REGION Network 5: State 2 = Valves Control
   RUNG wire#powerrail
      Contact( #RUNNING )
      { S7_Templates := "SrcType := Int" } GE_Contact(in1 := #STATE, in2 := 2)
      wire#w1
      { S7_Templates := "SrcType := Int" } LT_Contact(in1 := #STATE, in2 := 6)
      Coil( #OPN_AV )
   END_RUNG
   RUNG wire#w1
      { S7_Templates := "SrcType := Int" } LT_Contact(in1 := #STATE, in2 := 4)
      Coil( #OPN_FV1 )
   END_RUNG
   RUNG wire#w1
      { S7_Templates := "SrcType := Int" } LT_Contact(in1 := #STATE, in2 := 5)
      wire#w2
      Coil( #OPN_3W_FV2 )
   END_RUNG
   RUNG wire#w1
      { S7_Templates := "SrcType := Int" } GE_Contact(in1 := #STATE, in2 := 7)
      { S7_Templates := "SrcType := Int" } LE_Contact(in1 := #STATE, in2 := 8)
   END_RUNG wire#w2
   // the same network as SCL:
   #_w1 := #RUNNING AND (#STATE >= 2);
   #OPN_AV := #_w1 AND (#STATE < 6);
   #OPN_FV1 := #_w1 AND (#STATE < 4);
   #OPN_3W_FV2 := #_w1 AND ((#STATE < 5) OR ((#STATE >= 7) AND (#STATE <= 8)));
END_REGION

REGION Network 6: Into State 3
   RUNG wire#powerrail
      Contact( #RUNNING )
      { S7_Templates := "SrcType := Int" } EQ_Contact(in1 := #STATE, in2 := 2)
      Contact( #AV_Q )
      Contact( #FV1_Q )
      Contact( #FV2_3W_Q )
      Move(in := 3, out1 => #STATE)
   END_RUNG
   // the same network as SCL:
   IF #RUNNING AND (#STATE = 2) AND #AV_Q AND #FV1_Q AND #FV2_3W_Q THEN #STATE := 3; END_IF;
END_REGION

REGION Network 7: State 3 = Purge Active
   RUNG wire#powerrail
      Contact( #RUNNING )
      { S7_Templates := "SrcType := Int" } GE_Contact(in1 := #STATE, in2 := 3)
      { S7_Templates := "SrcType := Int" } LE_Contact(in1 := #STATE, in2 := 8)
      wire#w1
      Coil( #PRG_ACTV )
   END_RUNG
   RUNG wire#w1
      Coil( #ACTIVE )
   END_RUNG
   // the same network as SCL:
   #PRG_ACTV := #RUNNING AND (#STATE >= 3) AND (#STATE <= 8);
   #ACTIVE := #PRG_ACTV;
END_REGION

REGION Network 8: Into State 4
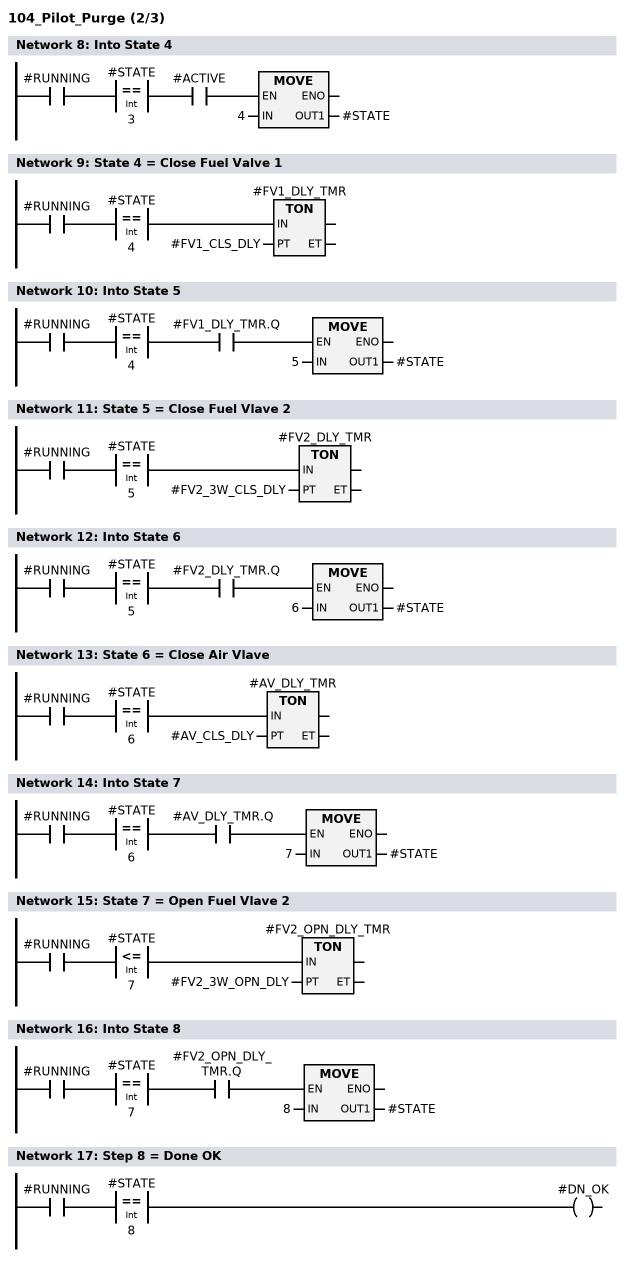
   RUNG wire#powerrail
      Contact( #RUNNING )
      { S7_Templates := "SrcType := Int" } EQ_Contact(in1 := #STATE, in2 := 3)
      Contact( #ACTIVE )
      Move(in := 4, out1 => #STATE)
   END_RUNG
   // the same network as SCL:
   IF #RUNNING AND (#STATE = 3) AND #ACTIVE THEN #STATE := 4; END_IF;
END_REGION

REGION Network 9: State 4 = Close Fuel Valve 1
   #FV1_DLY_TMR(IN := #RUNNING AND (#STATE = 4), PT := #FV1_CLS_DLY);   // TON
END_REGION

REGION Network 10: Into State 5
   RUNG wire#powerrail
      Contact( #RUNNING )
      { S7_Templates := "SrcType := Int" } EQ_Contact(in1 := #STATE, in2 := 4)
      Contact( #FV1_DLY_TMR.Q )
      Move(in := 5, out1 => #STATE)
   END_RUNG
   // the same network as SCL:
   IF #RUNNING AND (#STATE = 4) AND #FV1_DLY_TMR.Q THEN #STATE := 5; END_IF;
END_REGION

REGION Network 11: State 5 = Close Fuel Vlave 2
   #FV2_DLY_TMR(IN := #RUNNING AND (#STATE = 5), PT := #FV2_3W_CLS_DLY);   // TON
END_REGION

REGION Network 12: Into State 6
   RUNG wire#powerrail
      Contact( #RUNNING )
      { S7_Templates := "SrcType := Int" } EQ_Contact(in1 := #STATE, in2 := 5)
      Contact( #FV2_DLY_TMR.Q )
      Move(in := 6, out1 => #STATE)
   END_RUNG
   // the same network as SCL:
   IF #RUNNING AND (#STATE = 5) AND #FV2_DLY_TMR.Q THEN #STATE := 6; END_IF;
END_REGION

REGION Network 13: State 6 = Close Air Vlave
   #AV_DLY_TMR(IN := #RUNNING AND (#STATE = 6), PT := #AV_CLS_DLY);   // TON
END_REGION

REGION Network 14: Into State 7
   RUNG wire#powerrail
      Contact( #RUNNING )
      { S7_Templates := "SrcType := Int" } EQ_Contact(in1 := #STATE, in2 := 6)
      Contact( #AV_DLY_TMR.Q )
      Move(in := 7, out1 => #STATE)
   END_RUNG
   // the same network as SCL:
   IF #RUNNING AND (#STATE = 6) AND #AV_DLY_TMR.Q THEN #STATE := 7; END_IF;
END_REGION

REGION Network 15: State 7 = Open Fuel Vlave 2
   #FV2_OPN_DLY_TMR(IN := #RUNNING AND (#STATE <= 7), PT := #FV2_3W_OPN_DLY);   // TON
END_REGION

REGION Network 16: Into State 8
   RUNG wire#powerrail
      Contact( #RUNNING )
      { S7_Templates := "SrcType := Int" } EQ_Contact(in1 := #STATE, in2 := 7)
      Contact( #FV2_OPN_DLY_TMR.Q )
      Move(in := 8, out1 => #STATE)
   END_RUNG
   // the same network as SCL:
   IF #RUNNING AND (#STATE = 7) AND #FV2_OPN_DLY_TMR.Q THEN #STATE := 8; END_IF;
END_REGION

REGION Network 17: Step 8 = Done OK
   RUNG wire#powerrail
      Contact( #RUNNING )
      { S7_Templates := "SrcType := Int" } EQ_Contact(in1 := #STATE, in2 := 8)
      Coil( #DN_OK )
   END_RUNG
   // the same network as SCL:
   #DN_OK := #RUNNING AND (#STATE = 8);
END_REGION

REGION Network 18: Maximum Sequence Run Time
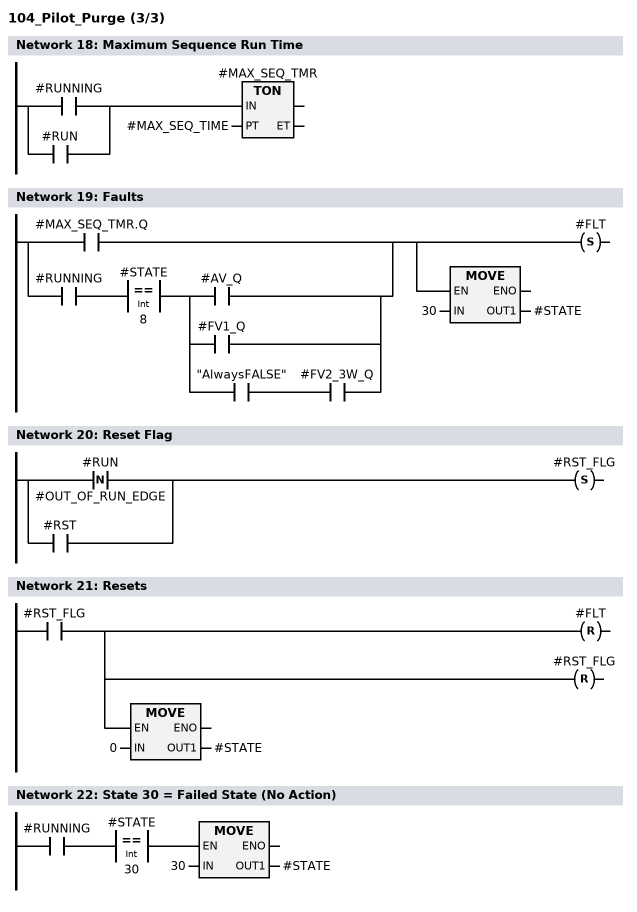
   #MAX_SEQ_TMR(IN := #RUNNING OR #RUN, PT := #MAX_SEQ_TIME);   // TON
END_REGION

REGION Network 19: Faults
   RUNG wire#powerrail
      Contact( #MAX_SEQ_TMR.Q )
      wire#w1
      S_Coil( #FLT )
   END_RUNG
   RUNG wire#powerrail
      Contact( #RUNNING )
      { S7_Templates := "SrcType := Int" } EQ_Contact(in1 := #STATE, in2 := 8)
      wire#w2
      Contact( #AV_Q )
   END_RUNG wire#w1
   RUNG wire#w2
      Contact( #FV1_Q )
   END_RUNG wire#w1
   RUNG wire#w2
      Contact( "AlwaysFALSE" )
      Contact( #FV2_3W_Q )
   END_RUNG wire#w1
   RUNG wire#w1
      Move(in := 30, out1 => #STATE)
   END_RUNG
   // the same network as SCL:
   IF #MAX_SEQ_TMR.Q OR (#RUNNING AND (#STATE = 8) AND (#AV_Q OR #FV1_Q OR ("AlwaysFALSE" AND #FV2_3W_Q))) THEN
       #FLT := TRUE;
       #STATE := 30;
   END_IF;
END_REGION

REGION Network 20: Reset Flag
   RUNG wire#powerrail
      N_Contact(operand := #RUN, bit := #OUT_OF_RUN_EDGE)
      wire#w1
      S_Coil( #RST_FLG )
   END_RUNG
   RUNG wire#powerrail
      Contact( #RST )
   END_RUNG wire#w1
   // the same network as SCL:
   #_w1 := NOT #RUN AND #OUT_OF_RUN_EDGE;   // falling edge of #RUN
   #OUT_OF_RUN_EDGE := #RUN;
   IF #_w1 OR #RST THEN #RST_FLG := TRUE; END_IF;
END_REGION

REGION Network 21: Resets
   RUNG wire#powerrail
      Contact( #RST_FLG )
      wire#w1
      R_Coil( #FLT )
   END_RUNG
   RUNG wire#w1
      R_Coil( #RST_FLG )
   END_RUNG
   RUNG wire#w1
      Move(in := 0, out1 => #STATE)
   END_RUNG
   // the same network as SCL:
   IF #RST_FLG THEN #FLT := FALSE; END_IF;
   #_w1 := #RST_FLG;
   IF #_w1 THEN
       #RST_FLG := FALSE;
       #STATE := 0;
   END_IF;
END_REGION

REGION Network 22: State 30 = Failed State (No Action)
   RUNG wire#powerrail
      Contact( #RUNNING )
      { S7_Templates := "SrcType := Int" } EQ_Contact(in1 := #STATE, in2 := 30)
      Move(in := 30, out1 => #STATE)
   END_RUNG
   // the same network as SCL:
   IF #RUNNING AND (#STATE = 30) THEN #STATE := 30; END_IF;
END_REGION
END_FUNCTION_BLOCK

FUNCTION_BLOCK "Evolving Setpoint"   // FB105, LAD
{ S7_Optimized_Access := 'TRUE' }
VERSION : 0.1
   VAR_INPUT
      Enable : Bool;
      Value : Real;
      Setpoint : Real;
      Gain : Real;
      Level_High : Real;
      Level_Low : Real;
   END_VAR
   VAR_OUTPUT
      Gain_Derived : Real;
      LevelBetter : Bool;
   END_VAR
   VAR
      "OFF Time" : TON_TIME;
      "On Time" : TON_TIME;
      Aux : Struct
         Aux_Derived : Bool;
         AuxSenzorDerivata1 : Real;
         AuxSenzorDerivata2 : Real;
         AuxSenzorDerivata11 : Real;
         AuxSenzorDerivata12 : Real;
         Puls_1 : Bool;
         Puls_2 : Bool;
         Puls_3 : Bool;
         Puls_4 : Bool;
         Gain_1 : Real;
      END_STRUCT;
      "Delay TOF" : TOF_TIME;
      "LevelBetter Delay" : TOF_TIME;
      "LevelBetter Prolong" : TOF_TIME;
   END_VAR
   VAR_TEMP   // added for the SCL form of the ladder/FBD networks
      _w1 : Bool;
      _w2 : Bool;
      _w3 : Bool;
      _w4 : Bool;
      _w5 : Bool;
      _w6 : Bool;
   END_VAR
BEGIN

REGION Network 1: Calcul derivata
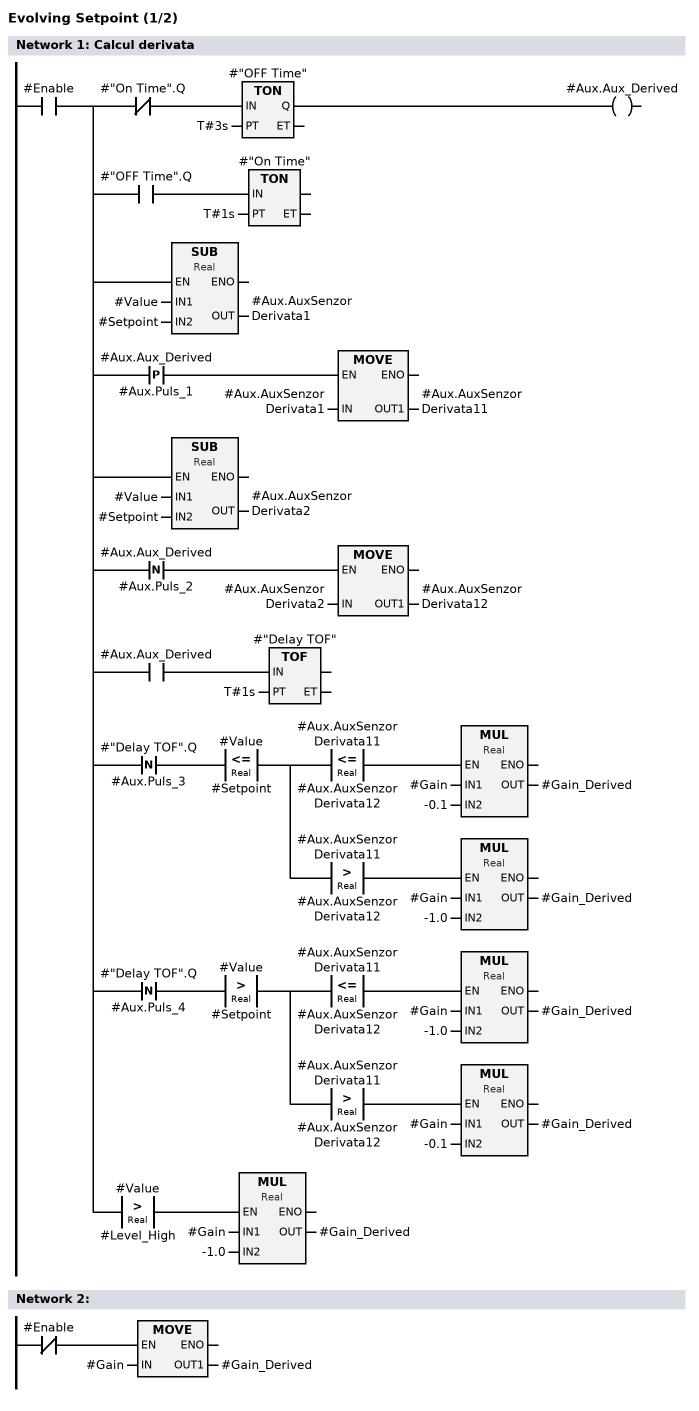
   #"OFF Time"(IN := #Enable AND NOT #"On Time".Q, PT := T#3s);   // TON
   #Aux.Aux_Derived := #"OFF Time".Q;
   #"On Time"(IN := #Enable AND #"OFF Time".Q, PT := T#1s);   // TON
   IF #Enable THEN #Aux.AuxSenzorDerivata1 := #Value - #Setpoint; END_IF;
   #_w1 := #Enable AND #Aux.Aux_Derived AND NOT #Aux.Puls_1;   // rising edge of #Aux.Aux_Derived
   #Aux.Puls_1 := #Aux.Aux_Derived;
   IF #_w1 THEN #Aux.AuxSenzorDerivata11 := #Aux.AuxSenzorDerivata1; END_IF;
   IF #Enable THEN #Aux.AuxSenzorDerivata2 := #Value - #Setpoint; END_IF;
   #_w2 := #Enable AND NOT #Aux.Aux_Derived AND #Aux.Puls_2;   // falling edge of #Aux.Aux_Derived
   #Aux.Puls_2 := #Aux.Aux_Derived;
   IF #_w2 THEN #Aux.AuxSenzorDerivata12 := #Aux.AuxSenzorDerivata2; END_IF;
   #"Delay TOF"(IN := #Enable AND #Aux.Aux_Derived, PT := T#1s);   // TOF
   #_w3 := #Enable AND NOT #"Delay TOF".Q AND #Aux.Puls_3;   // falling edge of #"Delay TOF".Q
   #Aux.Puls_3 := #"Delay TOF".Q;
   #_w4 := #_w3 AND (#Value <= #Setpoint);
   IF #_w4 AND (#Aux.AuxSenzorDerivata11 <= #Aux.AuxSenzorDerivata12) THEN
       #Gain_Derived := #Gain * (-0.1);
   END_IF;
   IF #_w4 AND (#Aux.AuxSenzorDerivata11 > #Aux.AuxSenzorDerivata12) THEN
       #Gain_Derived := #Gain * (-1.0);
   END_IF;
   #_w5 := #Enable AND NOT #"Delay TOF".Q AND #Aux.Puls_4;   // falling edge of #"Delay TOF".Q
   #Aux.Puls_4 := #"Delay TOF".Q;
   #_w6 := #_w5 AND (#Value > #Setpoint);
   IF #_w6 AND (#Aux.AuxSenzorDerivata11 <= #Aux.AuxSenzorDerivata12) THEN
       #Gain_Derived := #Gain * (-1.0);
   END_IF;
   IF #_w6 AND (#Aux.AuxSenzorDerivata11 > #Aux.AuxSenzorDerivata12) THEN
       #Gain_Derived := #Gain * (-0.1);
   END_IF;
   IF #Enable AND (#Value > #Level_High) THEN #Gain_Derived := #Gain * (-1.0); END_IF;
END_REGION

REGION Network 2
   RUNG wire#powerrail
      I_Contact( #Enable )
      { S7_GenerateENO := "TRUE" } Move(in := #Gain, out1 => #Gain_Derived)
   END_RUNG
   // the same network as SCL:
   IF NOT #Enable THEN #Gain_Derived := #Gain; END_IF;
END_REGION

REGION Network 3: Neautorizare pompa la imbunatatirea nivelului
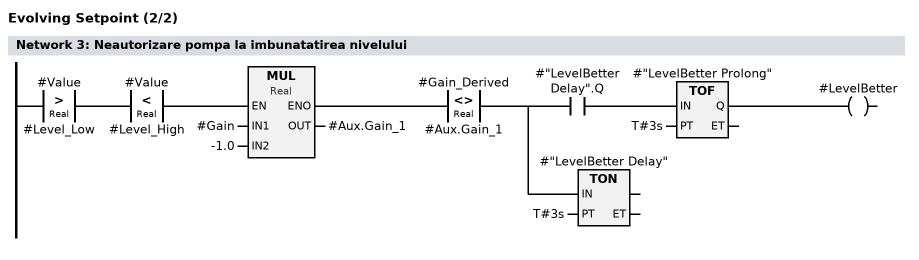
   // ENO of a box is taken as its EN; it also drops when the box reports an error
   #_w1 := (#Value > #Level_Low) AND (#Value < #Level_High);
   IF #_w1 THEN #Aux.Gain_1 := #Gain * (-1.0); END_IF;
   #_w2 := #_w1 AND (#Gain_Derived <> #Aux.Gain_1);
   #"LevelBetter Prolong"(IN := #_w2 AND #"LevelBetter Delay".Q, PT := T#3s);   // TOF
   #LevelBetter := #"LevelBetter Prolong".Q;
   #"LevelBetter Delay"(IN := #_w2, PT := T#3s);   // TON
END_REGION
END_FUNCTION_BLOCK

FUNCTION_BLOCK "106_O2_RAMP_CNTRL"   // FB106, LAD
TITLE = O2 Content Control Ramp
{ S7_Optimized_Access := 'TRUE' }
AUTHOR : JRS
VERSION : 0.1
// For the control of fuel pressure to maintain O2 level to specification
   VAR_INPUT
      RUN : Bool;   // Runs the block
      O2 : Real;   // Measured O2 level
      CBM : Bool;   // 1 = Cargo Blanketting Mode, 0 = Not
      BWT_SP : Real;   // BWT Setpoint
      CBM_SP : Real;   // CBM Setpoint
      CHK_TIME : Time;   // O2 Check delay from change
      RST : Bool;   // Reset bit
   END_VAR
   VAR_OUTPUT
      VLV_CNTRL : Real;   // Output to valve
   END_VAR
   VAR_IN_OUT
      RUNNING : Bool;   // Block is running
      INIT_CTRL_VAL : Real;   // Initial control value from modulation
   END_VAR
   VAR
      State : Int;   // State value for sequencing
      INTO_RUN_EDGE : Bool;   // Edge detection
      OUT_OF_RUN_EDGE : Bool;   // Edge detection
      RST_FLG : Bool;   // Reset flag
      VLV_DMND : Real;   // Valve demand value
      BIG_STEP : Real;   // Big change value
      MED_STEP : Real;   // Medium change value
      SML_STEP : Real;   // Small change value
      DISTANCE : Real;   // Distance to setpoint
      BIG_DIST : Real;   // Big distance
      MED_DIST : Real;   // Medium distance
      SML_DIST : Real;   // Small distance
      MEAS_DLY : TON_TIME;   // Measurement delay
      SETUP_DLY : TON_TIME;   // Setup delay
      CALC_DLY : TON_TIME;   // Calculation delay
      IEC_Timer_0_Instance : TP_TIME;
      IEC_Timer_0_Instance_1 : TON_TIME;
      "CALC_DLY 2" : TON_TIME;
      IEC_Timer_0_Instance_2 : TP_TIME;
      "Reset Sequence" : Bool;
      "Reset Sequence TP" : TP_TIME;
      IEC_Timer_0_Instance_3 : TON_TIME;
   END_VAR
   VAR_TEMP   // added for the SCL form of the ladder/FBD networks
      _w1 : Bool;
      _w2 : Bool;
      _w3 : Bool;
   END_VAR
BEGIN

REGION Network 1: Running
   // For running status detection
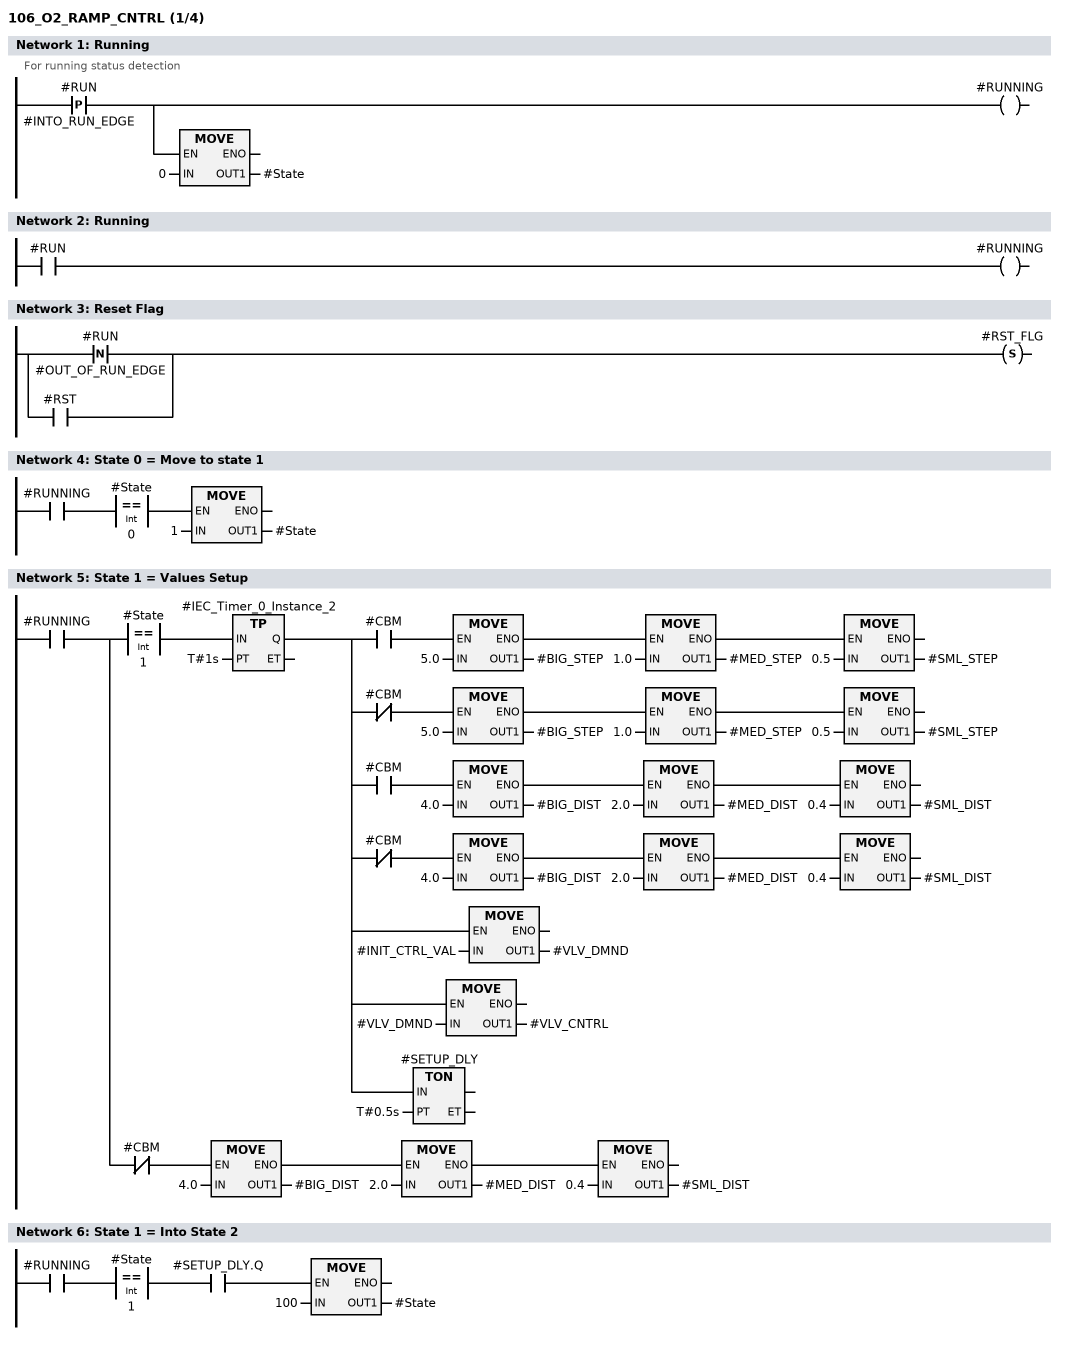
   RUNG wire#powerrail
      P_Contact(operand := #RUN, bit := #INTO_RUN_EDGE)
      wire#w1
      Coil( #RUNNING )
   END_RUNG
   RUNG wire#w1
      Move(in := 0, out1 => #State)
   END_RUNG
   // the same network as SCL:
   #_w1 := #RUN AND NOT #INTO_RUN_EDGE;   // rising edge of #RUN
   #INTO_RUN_EDGE := #RUN;
   #RUNNING := #_w1;
   IF #_w1 THEN #State := 0; END_IF;
END_REGION

REGION Network 2: Running
   RUNG wire#powerrail
      Contact( #RUN )
      Coil( #RUNNING )
   END_RUNG
   // the same network as SCL:
   #RUNNING := #RUN;
END_REGION

REGION Network 3: Reset Flag
   RUNG wire#powerrail
      N_Contact(operand := #RUN, bit := #OUT_OF_RUN_EDGE)
      wire#w1
      S_Coil( #RST_FLG )
   END_RUNG
   RUNG wire#powerrail
      Contact( #RST )
   END_RUNG wire#w1
   // the same network as SCL:
   #_w1 := NOT #RUN AND #OUT_OF_RUN_EDGE;   // falling edge of #RUN
   #OUT_OF_RUN_EDGE := #RUN;
   IF #_w1 OR #RST THEN #RST_FLG := TRUE; END_IF;
END_REGION

REGION Network 4: State 0 = Move to state 1
   RUNG wire#powerrail
      Contact( #RUNNING )
      { S7_Templates := "SrcType := Int" } EQ_Contact(in1 := #State, in2 := 0)
      Move(in := 1, out1 => #State)
   END_RUNG
   // the same network as SCL:
   IF #RUNNING AND (#State = 0) THEN #State := 1; END_IF;
END_REGION

REGION Network 5: State 1 = Values Setup
   #IEC_Timer_0_Instance_2(IN := #RUNNING AND (#State = 1), PT := T#1s);   // TP
   IF #IEC_Timer_0_Instance_2.Q AND #CBM THEN
       #BIG_STEP := 5.0;
       #MED_STEP := 1.0;
       #SML_STEP := 0.5;
   END_IF;
   IF #IEC_Timer_0_Instance_2.Q AND NOT #CBM THEN
       #BIG_STEP := 5.0;
       #MED_STEP := 1.0;
       #SML_STEP := 0.5;
   END_IF;
   IF #IEC_Timer_0_Instance_2.Q AND #CBM THEN
       #BIG_DIST := 4.0;
       #MED_DIST := 2.0;
       #SML_DIST := 0.4;
   END_IF;
   IF #IEC_Timer_0_Instance_2.Q AND NOT #CBM THEN
       #BIG_DIST := 4.0;
       #MED_DIST := 2.0;
       #SML_DIST := 0.4;
   END_IF;
   IF #IEC_Timer_0_Instance_2.Q THEN
       #VLV_DMND := #INIT_CTRL_VAL;
       #VLV_CNTRL := #VLV_DMND;
   END_IF;
   #SETUP_DLY(IN := #IEC_Timer_0_Instance_2.Q, PT := T#0.5s);   // TON
   IF #RUNNING AND NOT #CBM THEN
       #BIG_DIST := 4.0;
       #MED_DIST := 2.0;
       #SML_DIST := 0.4;
   END_IF;
END_REGION

REGION Network 6: State 1 = Into State 2
   RUNG wire#powerrail
      Contact( #RUNNING )
      { S7_Templates := "SrcType := Int" } EQ_Contact(in1 := #State, in2 := 1)
      Contact( #SETUP_DLY.Q )
      Move(in := 100, out1 => #State)
   END_RUNG
   // the same network as SCL:
   IF #RUNNING AND (#State = 1) AND #SETUP_DLY.Q THEN #State := 100; END_IF;
END_REGION

REGION Network 7: State 100 = Sequence reset
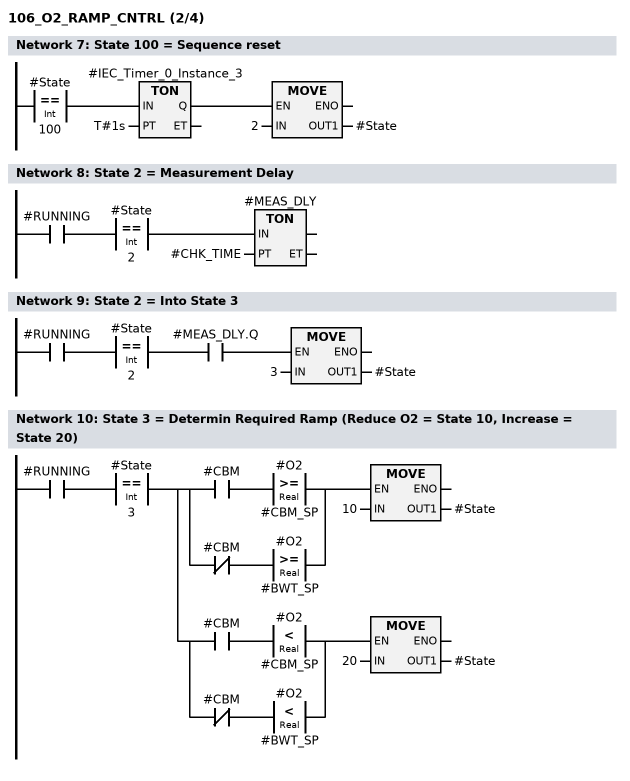
   #IEC_Timer_0_Instance_3(IN := #State = 100, PT := T#1s);   // TON
   IF #IEC_Timer_0_Instance_3.Q THEN #State := 2; END_IF;
END_REGION

REGION Network 8: State 2 = Measurement Delay
   #MEAS_DLY(IN := #RUNNING AND (#State = 2), PT := #CHK_TIME);   // TON
END_REGION

REGION Network 9: State 2 = Into State 3
   RUNG wire#powerrail
      Contact( #RUNNING )
      { S7_Templates := "SrcType := Int" } EQ_Contact(in1 := #State, in2 := 2)
      Contact( #MEAS_DLY.Q )
      Move(in := 3, out1 => #State)
   END_RUNG
   // the same network as SCL:
   IF #RUNNING AND (#State = 2) AND #MEAS_DLY.Q THEN #State := 3; END_IF;
END_REGION

REGION Network 10: State 3 = Determin Required Ramp (Reduce O2 = State 10, Increase = State 20)
   RUNG wire#powerrail
      Contact( #RUNNING )
      { S7_Templates := "SrcType := Int" } EQ_Contact(in1 := #State, in2 := 3)
      wire#w1
      Contact( #CBM )
      { S7_Templates := "SrcType := Real" } GE_Contact(in1 := #O2, in2 := #CBM_SP)
      wire#w2
      Move(in := 10, out1 => #State)
   END_RUNG
   RUNG wire#w1
      I_Contact( #CBM )
      { S7_Templates := "SrcType := Real" } GE_Contact(in1 := #O2, in2 := #BWT_SP)
   END_RUNG wire#w2
   RUNG wire#w1
      Contact( #CBM )
      { S7_Templates := "SrcType := Real" } LT_Contact(in1 := #O2, in2 := #CBM_SP)
      wire#w3
      Move(in := 20, out1 => #State)
   END_RUNG
   RUNG wire#w1
      I_Contact( #CBM )
      { S7_Templates := "SrcType := Real" } LT_Contact(in1 := #O2, in2 := #BWT_SP)
   END_RUNG wire#w3
   // the same network as SCL:
   #_w1 := #RUNNING AND (#State = 3);
   IF #_w1 AND ((#CBM AND (#O2 >= #CBM_SP)) OR (NOT #CBM AND (#O2 >= #BWT_SP))) THEN #State := 10; END_IF;
   IF #_w1 AND ((#CBM AND (#O2 < #CBM_SP)) OR (NOT #CBM AND (#O2 < #BWT_SP))) THEN #State := 20; END_IF;
END_REGION

REGION Network 12: State 10 = Reduce O2 = Increase Fuel Pressure = Open Valve (Calculations)
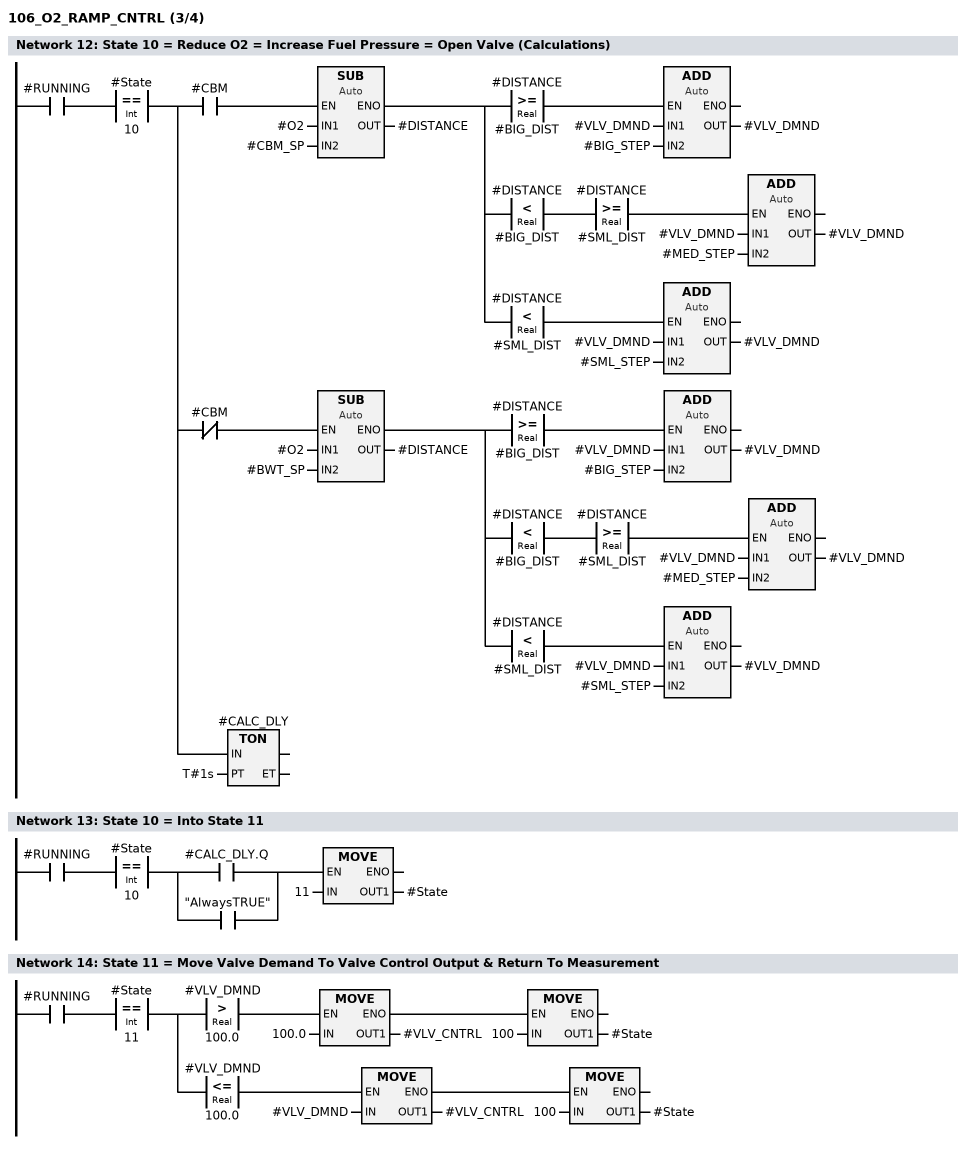
   #_w1 := #RUNNING AND (#State = 10);
   #_w2 := #_w1 AND #CBM;
   IF #_w2 THEN #DISTANCE := #O2 - #CBM_SP; END_IF;
   IF #_w2 AND (#DISTANCE >= #BIG_DIST) THEN #VLV_DMND := #VLV_DMND + #BIG_STEP; END_IF;
   IF #_w2 AND (#DISTANCE < #BIG_DIST) AND (#DISTANCE >= #SML_DIST) THEN
       #VLV_DMND := #VLV_DMND + #MED_STEP;
   END_IF;
   IF #_w2 AND (#DISTANCE < #SML_DIST) THEN #VLV_DMND := #VLV_DMND + #SML_STEP; END_IF;
   #_w3 := #_w1 AND NOT #CBM;
   IF #_w3 THEN #DISTANCE := #O2 - #BWT_SP; END_IF;
   IF #_w3 AND (#DISTANCE >= #BIG_DIST) THEN #VLV_DMND := #VLV_DMND + #BIG_STEP; END_IF;
   IF #_w3 AND (#DISTANCE < #BIG_DIST) AND (#DISTANCE >= #SML_DIST) THEN
       #VLV_DMND := #VLV_DMND + #MED_STEP;
   END_IF;
   IF #_w3 AND (#DISTANCE < #SML_DIST) THEN #VLV_DMND := #VLV_DMND + #SML_STEP; END_IF;
   #CALC_DLY(IN := #_w1, PT := T#1s);   // TON
END_REGION

REGION Network 13: State 10 = Into State 11
   RUNG wire#powerrail
      Contact( #RUNNING )
      { S7_Templates := "SrcType := Int" } EQ_Contact(in1 := #State, in2 := 10)
      wire#w1
      Contact( #CALC_DLY.Q )
      wire#w2
      Move(in := 11, out1 => #State)
   END_RUNG
   RUNG wire#w1
      Contact( "AlwaysTRUE" )
   END_RUNG wire#w2
   // the same network as SCL:
   IF #RUNNING AND (#State = 10) AND (#CALC_DLY.Q OR "AlwaysTRUE") THEN #State := 11; END_IF;
END_REGION

REGION Network 14: State 11 = Move Valve Demand To Valve Control Output & Return To Measurement
   RUNG wire#powerrail
      Contact( #RUNNING )
      { S7_Templates := "SrcType := Int" } EQ_Contact(in1 := #State, in2 := 11)
      wire#w1
      { S7_Templates := "SrcType := Real" } GT_Contact(in1 := #VLV_DMND, in2 := 100.0)
      Move(in := 100.0, out1 => #VLV_CNTRL)
      Move(in := 100, out1 => #State)
   END_RUNG
   RUNG wire#w1
      { S7_Templates := "SrcType := Real" } LE_Contact(in1 := #VLV_DMND, in2 := 100.0)
      Move(in := #VLV_DMND, out1 => #VLV_CNTRL)
      Move(in := 100, out1 => #State)
   END_RUNG
   // the same network as SCL:
   #_w1 := #RUNNING AND (#State = 11);
   IF #_w1 AND (#VLV_DMND > 100.0) THEN
       #VLV_CNTRL := 100.0;
       #State := 100;
   END_IF;
   IF #_w1 AND (#VLV_DMND <= 100.0) THEN
       #VLV_CNTRL := #VLV_DMND;
       #State := 100;
   END_IF;
END_REGION

REGION Network 16: State 20 = Increase O2 = Decrease Fuel Pressure = Close Valve (Calculations)
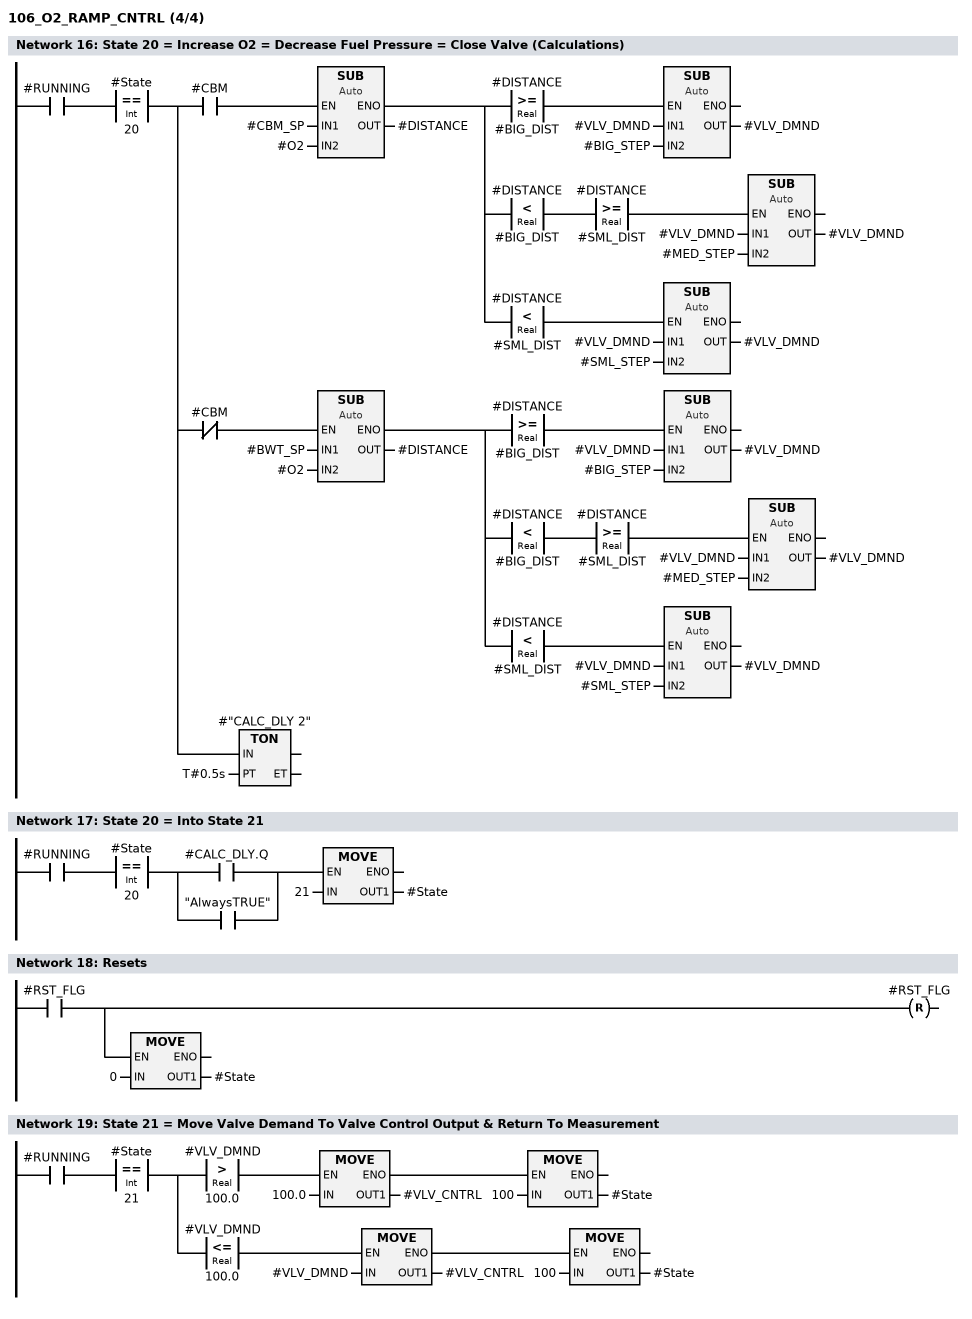
   #_w1 := #RUNNING AND (#State = 20);
   #_w2 := #_w1 AND #CBM;
   IF #_w2 THEN #DISTANCE := #CBM_SP - #O2; END_IF;
   IF #_w2 AND (#DISTANCE >= #BIG_DIST) THEN #VLV_DMND := #VLV_DMND - #BIG_STEP; END_IF;
   IF #_w2 AND (#DISTANCE < #BIG_DIST) AND (#DISTANCE >= #SML_DIST) THEN
       #VLV_DMND := #VLV_DMND - #MED_STEP;
   END_IF;
   IF #_w2 AND (#DISTANCE < #SML_DIST) THEN #VLV_DMND := #VLV_DMND - #SML_STEP; END_IF;
   #_w3 := #_w1 AND NOT #CBM;
   IF #_w3 THEN #DISTANCE := #BWT_SP - #O2; END_IF;
   IF #_w3 AND (#DISTANCE >= #BIG_DIST) THEN #VLV_DMND := #VLV_DMND - #BIG_STEP; END_IF;
   IF #_w3 AND (#DISTANCE < #BIG_DIST) AND (#DISTANCE >= #SML_DIST) THEN
       #VLV_DMND := #VLV_DMND - #MED_STEP;
   END_IF;
   IF #_w3 AND (#DISTANCE < #SML_DIST) THEN #VLV_DMND := #VLV_DMND - #SML_STEP; END_IF;
   #"CALC_DLY 2"(IN := #_w1, PT := T#0.5s);   // TON
END_REGION

REGION Network 17: State 20 = Into State 21
   RUNG wire#powerrail
      Contact( #RUNNING )
      { S7_Templates := "SrcType := Int" } EQ_Contact(in1 := #State, in2 := 20)
      wire#w1
      Contact( #CALC_DLY.Q )
      wire#w2
      Move(in := 21, out1 => #State)
   END_RUNG
   RUNG wire#w1
      Contact( "AlwaysTRUE" )
   END_RUNG wire#w2
   // the same network as SCL:
   IF #RUNNING AND (#State = 20) AND (#CALC_DLY.Q OR "AlwaysTRUE") THEN #State := 21; END_IF;
END_REGION

REGION Network 18: Resets
   RUNG wire#powerrail
      Contact( #RST_FLG )
      wire#w1
      R_Coil( #RST_FLG )
   END_RUNG
   RUNG wire#w1
      Move(in := 0, out1 => #State)
   END_RUNG
   // the same network as SCL:
   #_w1 := #RST_FLG;
   IF #_w1 THEN
       #RST_FLG := FALSE;
       #State := 0;
   END_IF;
END_REGION

REGION Network 19: State 21 = Move Valve Demand To Valve Control Output & Return To Measurement
   RUNG wire#powerrail
      Contact( #RUNNING )
      { S7_Templates := "SrcType := Int" } EQ_Contact(in1 := #State, in2 := 21)
      wire#w1
      { S7_Templates := "SrcType := Real" } GT_Contact(in1 := #VLV_DMND, in2 := 100.0)
      Move(in := 100.0, out1 => #VLV_CNTRL)
      Move(in := 100, out1 => #State)
   END_RUNG
   RUNG wire#w1
      { S7_Templates := "SrcType := Real" } LE_Contact(in1 := #VLV_DMND, in2 := 100.0)
      Move(in := #VLV_DMND, out1 => #VLV_CNTRL)
      Move(in := 100, out1 => #State)
   END_RUNG
   // the same network as SCL:
   #_w1 := #RUNNING AND (#State = 21);
   IF #_w1 AND (#VLV_DMND > 100.0) THEN
       #VLV_CNTRL := 100.0;
       #State := 100;
   END_IF;
   IF #_w1 AND (#VLV_DMND <= 100.0) THEN
       #VLV_CNTRL := #VLV_DMND;
       #State := 100;
   END_IF;
END_REGION
END_FUNCTION_BLOCK

FUNCTION "100_SC" : Void   // FC100, LAD
TITLE = State Complete
{ S7_Optimized_Access := 'TRUE' }
AUTHOR : JRS
VERSION : 0.1
// For the determination of each step state being complete
BEGIN

REGION Network 1: Step 001 = Confirm Auto Conditions Ok
